sDate := DateFormat(stTime:= fbGetTime.dtDateAndTime);
//----------------------------------------------------------------------------------------------
// Delete
//----------------------------------------------------------------------------------------------
IF rtDelete.Q THEN
	FOR uiI := 1 TO cuiSize DO
		IF astErrorEvent[uiI].sErrorID = sErrorID THEN
			SysMemMove(pSrc := ADR(astErrorEvent[uiI+1]), pDest := ADR(astErrorEvent[uiI]), udiCount :=  SIZEOF(st_ErrorEvent) * (cuiSize-uiI));
			astErrorEvent[cuiSize].sErrorID		:= 'No error';
			EXIT;		
		END_IF
	END_FOR
END_IF

END_FUNCTION_BLOCK

// Programs/Tools/DateFormat
FUNCTION DateFormat : STRING
VAR_INPUT
	///Time input from ErrorFifo
	stTime: DATE_AND_TIME;
END_VAR
VAR
	///Date output in string
	sDate : STRING;
	sTemp : STRING;
	sDateTime: STRING := '';
END_VAR

//------------------------------------------------------------------------
// To show the date in the errortable in a usable format
//------------------------------------------------------------------------	

sDate := DT_TO_STRING(stTime);

//------------------------------------------------------------------------
// Cutting the days
//------------------------------------------------------------------------	

sTemp := sDate;
sDateTime := MID(STR:= sTemp, LEN:= 2, POS:= 12);
sDateTime := CONCAT(sDateTime, '/');
	
//------------------------------------------------------------------------
// Cutting the months
//------------------------------------------------------------------------		
sTemp := sDate;
sDateTime := CONCAT(sDateTime, MID(STR:= sTemp, LEN:= 2, POS:= 9));
sDateTime := CONCAT(sDateTime, '/');

//------------------------------------------------------------------------
// Cutting the years
//------------------------------------------------------------------------		

sTemp := sDate;
sDateTime := CONCAT(sDateTime, MID(STR:= sTemp, LEN:= 4, POS:= 4));
sDateTime := CONCAT(sDateTime, ' - ');	
	
//------------------------------------------------------------------------
// Cutting the hours and minutes and seconds
//------------------------------------------------------------------------	

sTemp := sDate;
sDateTime := CONCAT(sDateTime, RIGHT(STR:= sTemp, SIZE:= 8)	);

//------------------------------------------------------------------------		


	DateFormat := sDateTime;

END_FUNCTION

// Programs/Tools/MovCntr2B2M
FUNCTION_BLOCK MovCntr2B2M
VAR_INPUT
	/// Flag to Reset Error
	xQuit: BOOL;
	/// Enable error reset flag
	xQuitEN: BOOL;
	/// Enable error control
	xEnable: BOOL;
	/// Limit switch for movement 1 (M1 <--> B1) 
	xB1: BOOL;
	/// Limit switch for movement 2 (M2 <--> B2) 
	xB2: BOOL;
	/// Actor Signal for movement 1 (M1 <--> B1) 
	xM1: BOOL;
	/// Actor Signal for movement 1 (M2 <--> B2) 
	xM2: BOOL;
	/// Timeout-Time for movement 1	
	T1: TIME;
	/// Timeout-Time for movement 2
	T2: TIME;
END_VAR
VAR
	/// Timeout timer for movement 1
	TON1: TON;
	/// Timeout timer for movement 2
	TON2: TON;
	/// SR FlipFlop for Err1
	RS1: RS;
	/// SR FlipFlop for Err2
	RS2: RS;
END_VAR
VAR_OUTPUT
	/// Timeout movement 1
	xErr1: BOOL;
	/// Timeout movement 2 
	xErr2: BOOL;
END_VAR

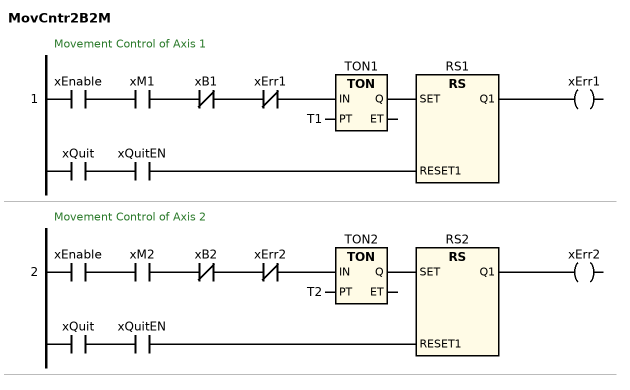
// NETWORK 1
// Movement Control of Axis 1
TON1(IN := xEnable AND xM1 AND NOT xB1 AND NOT xErr1, PT := T1); // TON
RS1(SET := TON1.Q, RESET1 := xQuit AND xQuitEN); // RS
xErr1 := RS1.Q1;

// NETWORK 2
// Movement Control of Axis 2
TON2(IN := xEnable AND xM2 AND NOT xB2 AND NOT xErr2, PT := T2); // TON
RS2(SET := TON2.Q, RESET1 := xQuit AND xQuitEN); // RS
xErr2 := RS2.Q1;

END_FUNCTION_BLOCK

// Programs/Visu/VisuProgramStp
PROGRAM  VisuProgramStp
VAR
	blBlink	: BLINK;
	t: TIME;
	uiNumOfApplications	: UINT:= 1;
	uiNumOfStoppers		: UINT:= 1;
	rtConvR				: R_TRIG;
	rtConvL				: R_TRIG;
	rtConvS				: R_TRIG;
	byActiveMainScreen	: BYTE;
	byActiveSubScreen	: BYTE;
	byScreenTitle		: BYTE;
	uiI					: UINT;
	astErrorEvents		: ARRAY [1..20] OF st_ErrorEvent;
	rtTime				: R_TRIG;
	fbGetTime: RTCLK.GetDateAndTime;
	sDate: STRING;
	dtTime	: DATE_AND_TIME;
	uiCarrierInitNum: UINT;
	xCarrierInit: BOOL;
	tonDefErr: TON;
	tonMesErr: TON;
	tonSapErr: TON;
	
	stRfidCdpx	: dc_ecp.st_CPF_RfidData;
	astAppControlONo: UDINT;
END_VAR

byActiveMainScreen	:= BOOL_TO_BYTE(fromCDPX.stCdpxButtonState.xHome)*0 + BOOL_TO_BYTE(fromCDPX.stCdpxButtonState.xSetupMode)*1 + BOOL_TO_BYTE(fromCDPX.stCdpxButtonState.xParameter)*2 + BOOL_TO_BYTE(fromCDPX.stCdpxButtonState.xSystem)*3;
byActiveSubScreen	:= BOOL_TO_BYTE(fromCDPX.stCdpxButtonState.xOperationMode)*0 + BOOL_TO_BYTE(fromCDPX.stCdpxButtonState.xApp_1)*0 +  BOOL_TO_BYTE(fromCDPX.stCdpxButtonState.xApp)*0 + BOOL_TO_BYTE(fromCDPX.stCdpxButtonState.xSystem)*0 + BOOL_TO_BYTE(fromCDPX.stCdpxButtonState.xOverview)*1 + BOOL_TO_BYTE(fromCDPX.stCdpxButtonState.xApp_2)*1 +  BOOL_TO_BYTE(fromCDPX.stCdpxButtonState.xTrans_1)*1 + BOOL_TO_BYTE(fromCDPX.stCdpxButtonState.xUser)*2 + BOOL_TO_BYTE(fromCDPX.stCdpxButtonState.xBelt)*2 +  BOOL_TO_BYTE(fromCDPX.stCdpxButtonState.xTrans_2)*2 + BOOL_TO_BYTE(fromCDPX.stCdpxButtonState.xStp_1)*3+ BOOL_TO_BYTE(fromCDPX.stCdpxButtonState.xStp_2)*4;
byScreenTitle 		:= byActiveMainScreen* 10 + byActiveSubScreen  ;

dtTime := fbGetTime.dtDateAndTime;
rtTime(CLK:= fbGetTime.xDone);
IF rtTime.Q THEN
sDate := DateFormat(stTime:= dtTime);
END_IF
fbGetTime( xExecute:= NOT fbGetTime.xDone);
fbGetTime( xExecute:= fbGetTime.xDone);

//////////////////////////////////
//			from CDPX			//
//////////////////////////////////

IF xFirstCycle THEN
	fromCDPX.astTransitionTable_1:= astTransitionTableStopper1 ;
	fromCDPX.uiMode := 1;
ELSE	
	astTransitionTableStopper1 :=fromCDPX.astTransitionTable_1;
	Visu.byMode 			:= UINT_TO_BYTE(fromCDPX.uiMode);
END_IF

// DABO /////////////////////////////////////////////////////////////////////////
IF uiCarrierInitNum <> stpStopper1.stAppSettings.uiCarrierInitNum THEN
	uiCarrierInitNum := stpStopper1.stAppSettings.uiCarrierInitNum;
ELSIF uiCarrierInitNum <> fromCDPX.astAppSetting[0].uiCarrierInitNum THEN
	uiCarrierInitNum := fromCDPX.astAppSetting[0].uiCarrierInitNum;
END_IF

fromCDPX.astAppSetting[0].uiCarrierInitNum := uiCarrierInitNum;
SysMemCpy(pDest:= ADR(stpStopper1.stAppSettings.uiCarrierInitNum), pSrc:= ADR(uiCarrierInitNum), udiCount:= SIZEOF(uiCarrierInitNum));

IF xCarrierInit <> stpStopper1.stAppSettings.xCarrierInit THEN
	xCarrierInit := stpStopper1.stAppSettings.xCarrierInit;
ELSIF xCarrierInit <> fromCDPX.astAppSetting[0].xCarrierInit THEN
	xCarrierInit := fromCDPX.astAppSetting[0].xCarrierInit;
END_IF

fromCDPX.astAppSetting[0].xCarrierInit := xCarrierInit;
SysMemCpy(pDest:= ADR(stpStopper1.stAppSettings.xCarrierInit), pSrc:= ADR(xCarrierInit), udiCount:= SIZEOF(xCarrierInit));

SysMemCpy(pDest:= ADR(stpStopper1.stAppSettings.xActive), pSrc:= ADR(fromCDPX.astAppSetting[0].xActive), udiCount:= SIZEOF(fromCDPX.astAppSetting[0].xActive));
SysMemCpy(pDest:= ADR(stpStopper1.stAppSettings.xStopBelt), pSrc:= ADR(fromCDPX.astAppSetting[0].xStopBelt), udiCount:= SIZEOF(fromCDPX.astAppSetting[0].xStopBelt));

//////////////////////////////////////////////////////////////////////////////////
// conveyor handling
rtConvL(CLK:= fromCDPX.astConveyorButtonState[0].xConvLeft);
rtConvR(CLK:= fromCDPX.astConveyorButtonState[0].xConvRight);
rtConvS(CLK:= fromCDPX.astConveyorButtonState[0].xConvSlow);
IF rtConvL.Q THEN
	IF  stpStopper1.convConveyor.xLeft THEN
		stpStopper1.convConveyor.Stop();
	ELSE
		stpStopper1.convConveyor.RunToLeft(stpStopper1.convConveyor.xSlow);
	END_IF
END_IF
IF rtConvR.Q THEN
	IF  stpStopper1.convConveyor.xRight THEN
		stpStopper1.convConveyor.Stop();
	ELSE
		stpStopper1.convConveyor.RunToRight(stpStopper1.convConveyor.xSlow);
	END_IF
END_IF
IF rtConvS.Q THEN
	IF  stpStopper1.convConveyor.xSlow THEN
		stpStopper1.convConveyor.SpeedUp();
	ELSE
		stpStopper1.convConveyor.SlowDown();
	END_IF
END_IF

// Operation mode buttons
fromCDPX.stHome_OperationMode_Reset.xActive := xReset OR (xResetEn AND blBlink.OUT);
fromCDPX.stHome_OperationMode_Reset.xDisabled := NOT xResetEn;

fromCDPX.stHome_OperationMode_Automatic.xActive := xAuto OR (xAutoEn AND blBlink.OUT);
fromCDPX.stHome_OperationMode_Automatic.xDisabled := NOT xAutoEn AND NOT xAuto;

fromCDPX.stHome_OperationMode_Setup.xActive := xManual;
fromCDPX.stHome_OperationMode_Setup.xDisabled := NOT xManualEn AND NOT xManual;

fromCDPX.stHome_OperationMode_CycleEnd.xActive := xCycleEnd AND blBlink.OUT;
fromCDPX.stHome_OperationMode_CycleEnd.xDisabled := NOT xCycleEndEn AND NOT xCycleEnd;

stWinCC.xAuto 		:= fromCDPX.stHome_OperationMode_Automatic.xPressed;
stWinCC.xReset 		:= fromCDPX.stHome_OperationMode_Reset.xPressed;
stWinCC.xManual 	:= fromCDPX.stHome_OperationMode_Setup.xPressed;
stWinCC.xCycleEnd 	:= fromCDPX.stHome_OperationMode_CycleEnd.xPressed;
stWinCC.xQuit		:= fromCDPX.stCdpxButtonState.xClearError;

// Setup RFID buttons
fromCDPX.stSetupMode_Stopper1_Init.xActive R= stpStopper1.stpStopper.dtmRfid.xReady;
fromCDPX.stSetupMode_Stopper1_Init.xActive S= fromCDPX.stSetupMode_Stopper1_Init.xPressed;
fromCDPX.stSetupMode_Stopper1_Init.xDisabled :=  xManual;
IF fromCDPX.astStopperButton[0].xInit THEN
	stpStopper1.stpStopper.Connect(usiCanChannel := stpStopper1.usiCanChannel, usiCanNetworkId := stpStopper1.usiCanNetworkId, usiCanNodeId := stpStopper1.usiCanNodeId);
END_IF


fromCDPX.stSetupMode_Stopper1_Read.xActive R= stpStopper1.stpStopper.dtmRfid.xReady;
fromCDPX.stSetupMode_Stopper1_Read.xActive S= fromCDPX.stSetupMode_Stopper1_Read.xPressed;
fromCDPX.stSetupMode_Stopper1_Read.xDisabled := xManual;
IF fromCDPX.astStopperButton[0].xRead THEN
	stpStopper1.stpStopper.ReadRfid(pstRfidData := ADR(stRfidCdpx));
	toCDPX.astRfidData[0].uiCarrierID				:=	stRfidCdpx.uiCarrierID					 ;
	toCDPX.astRfidData[0].uiCode					:=	stRfidCdpx.uiCode						 	;
	toCDPX.astRfidData[0].uiParameter1				:=	stRfidCdpx.uiParameter1					 ;
	toCDPX.astRfidData[0].uiParameter2				:=	stRfidCdpx.uiParameter2					 ;
	toCDPX.astRfidData[0].uiParameter3				:=	stRfidCdpx.uiParameter3					 ;
	toCDPX.astRfidData[0].uiParameter4				:=	stRfidCdpx.uiParameter4					 ;
	toCDPX.astRfidData[0].stMesData.udiONo			:=	stRfidCdpx.stMesData.udiONo				 ;
	toCDPX.astRfidData[0].stMesData.udiPNo			:=	stRfidCdpx.stMesData.udiPNo				 ;
	toCDPX.astRfidData[0].stMesData.uiOpNo			:=	stRfidCdpx.stMesData.uiOpNo				 ;
	toCDPX.astRfidData[0].stMesData.uiOPos			:=	stRfidCdpx.stMesData.uiOPos				 ;
	toCDPX.astRfidData[0].stMesData.uiResourceId	:=	stRfidCdpx.stMesData.uiResourceId		 	;
	toCDPX.astRfidData[0].stSapData.sItem	 		:=	stRfidCdpx.stSapData.sItem	 			 ;
	toCDPX.astRfidData[0].stSapData.sItemRev		:=	stRfidCdpx.stSapData.sItemRev			 	;
	toCDPX.astRfidData[0].stSapData.sSfc			:=	stRfidCdpx.stSapData.sSfc				 	;
	toCDPX.astRfidData[0].stSapData.udiOp			:=	stRfidCdpx.stSapData.udiOp				 ;
	toCDPX.astRfidData[0].stSapData.udiSfc			:=	stRfidCdpx.stSapData.udiSfc				 ;
END_IF                                                	


fromCDPX.stSetupMode_Stopper1_Write.xActive R= stpStopper1.stpStopper.dtmRfid.xReady;
fromCDPX.stSetupMode_Stopper1_Write.xActive S= fromCDPX.stSetupMode_Stopper1_Write.xPressed;
fromCDPX.stSetupMode_Stopper1_Write.xDisabled := xManual;
IF fromCDPX.astStopperButton[0].xWrite THEN
	stRfidCdpx.uiCarrierID					:= toCDPX.astRfidData[0].uiCarrierID				;
	stRfidCdpx.uiCode						:= toCDPX.astRfidData[0].uiCode					;
	stRfidCdpx.uiParameter1					:= toCDPX.astRfidData[0].uiParameter1				;
	stRfidCdpx.uiParameter2					:= toCDPX.astRfidData[0].uiParameter2				;
	stRfidCdpx.uiParameter3					:= toCDPX.astRfidData[0].uiParameter3				;
	stRfidCdpx.uiParameter4					:= toCDPX.astRfidData[0].uiParameter4				;
	stRfidCdpx.stMesData.udiONo				:= toCDPX.astRfidData[0].stMesData.udiONo			;
	stRfidCdpx.stMesData.udiPNo				:= toCDPX.astRfidData[0].stMesData.udiPNo			;
	stRfidCdpx.stMesData.uiOpNo				:= toCDPX.astRfidData[0].stMesData.uiOpNo			;
	stRfidCdpx.stMesData.uiOPos				:= toCDPX.astRfidData[0].stMesData.uiOPos			;
	stRfidCdpx.stMesData.uiResourceId		:= toCDPX.astRfidData[0].stMesData.uiResourceId	;
	stRfidCdpx.stSapData.sItem	 			:= toCDPX.astRfidData[0].stSapData.sItem	 		;
	stRfidCdpx.stSapData.sItemRev			:= toCDPX.astRfidData[0].stSapData.sItemRev		;
	stRfidCdpx.stSapData.sSfc				:= toCDPX.astRfidData[0].stSapData.sSfc			;
	stRfidCdpx.stSapData.udiOp				:= toCDPX.astRfidData[0].stSapData.udiOp			;
	stRfidCdpx.stSapData.udiSfc				:= toCDPX.astRfidData[0].stSapData.udiSfc			;
	stpStopper1.stpStopper.WriteRfid(stRfidData:= stRfidCdpx);
END_IF


fromCDPX.stSetupMode_Stopper1_DeleteData.xActive := fromCDPX.stSetupMode_Stopper1_DeleteData.xPressed;
fromCDPX.stSetupMode_Stopper1_DeleteData.xDisabled := xManual;                                            
IF fromCDPX.astStopperButton[0].xDeleteData	THEN
	SysMemSet(pDest:= ADR(stpStopper1.stpStopper.stRfidVisu), udiValue:= 0, udiCount:= SIZEOF(stpStopper1.stpStopper.stRfidVisu));
	SysMemCpy(pDest:= ADR(toCDPX.astRfidData[0]), pSrc:= ADR(stpStopper1.stpStopper.stRfidVisu), udiCount:= SIZEOF(stpStopper1.stpStopper.stRfidData));	
END_IF

IF NOt xManual  THEN
	SysMemCpy(pDest:= ADR(toCDPX.astRfidData[0]), pSrc:= ADR(stpStopper1.stpStopper.stRfidVisu), udiCount:= SIZEOF(stpStopper1.stpStopper.stRfidData));	
END_IF


IF fromCDPX.astStopperButton[0].xStpMveDown	THEN
	stpStopper1.stpStopper.cpfssStopper.StayDown();
END_IF
IF fromCDPX.astStopperButton[0].xStpMveUp	THEN
	stpStopper1.stpStopper.cpfssStopper.MoveUp();
END_IF

Visu.stInteractiveError.xBtnAbort 		:= fromCDPX.stInteractiveMessage_Abort.xPressed;
Visu.stInteractiveError.xBtnIgnore 		:= fromCDPX.stInteractiveMessage_Ignore.xPressed;
Visu.stInteractiveError.xBtnRejectOrder := fromCDPX.stInteractiveMessage_RejectOrder.xPressed;
Visu.stInteractiveError.xBtnRepeat		:= fromCDPX.stInteractiveMessage_Repeat.xPressed;

blBlink(ENABLE := TRUE, TIMEHIGH := T#1S, TIMELOW := T#1S); 
	

IF Visu.byMode = 1 THEN
	xMES := TRUE;
	xSAP := FALSE;
ELSIF Visu.byMode = 2 THEN
	xMES := FALSE;
	xSAP := TRUE;
ELSE
	xMES := FALSE;
	xSAP := FALSE;
END_IF

IF NOT xAuto AND NOT xManual AND NOT xReset THEN
	Visu.byOpMode := 0;
ELSIF xReset THEN
	Visu.byOpMode := 1;
ELSIF xAuto THEN
	Visu.byOpMode := 2;
ELSIF xManual THEN
	Visu.byOpMode := 3;
END_IF


//////////////////////////////////
//			to CDPX				//
//////////////////////////////////


toCDPX.byOpMode									:= Visu.byOpMode;
toCDPX.byScreenTitle							:= byScreenTitle;
toCDPX.xManual									:= xManual;	
toCDPX.xAuto									:= xAuto;			
toCDPX.xSAP										:= xSAP;				
toCDPX.xMES										:= xMES;				
toCDPX.xDefault									:= NOT xSAP AND NOT xMES;		
toCDPX.uiNumOfApplications						:= uiNumOfApplications;				
toCDPX.uiNumOfStoppers							:= uiNumOfStoppers;						
toCDPX.sDate									:= LEFT(sDate,10);
toCDPX.sTime									:= RIGHT(sDate,8);
toCDPX.auiCondIn[0]								:= stpStopper1.uiCondIn;
toCDPX.auiCondOut[0]							:= stpStopper1.uiCondOut;


toCDPX.astSensorSignals[0].sInductive_1			:= 'xBG21';
toCDPX.astSensorSignals[0].sInductive_2			:= 'xBG22';
toCDPX.astSensorSignals[0].sInductive_3			:= 'xBG23';
toCDPX.astSensorSignals[0].sInductive_4			:= 'xBG24';
toCDPX.astSensorSignals[0].sRfid				:= 'TF80';
toCDPX.astSensorSignals[0].sStpDownOutpu		:= 'xMB20';
toCDPX.astSensorSignals[0].sStpDownSensor		:= 'xBG20';
toCDPX.astSensorSignals[0].xInductive_1			:= xBG21; 
toCDPX.astSensorSignals[0].xInductive_2			:= xBG22; 
toCDPX.astSensorSignals[0].xInductive_3			:= xBG23; 
toCDPX.astSensorSignals[0].xInductive_4			:= xBG24; 
toCDPX.astSensorSignals[0].xStpDownOutpu		:= xMB20; 
toCDPX.astSensorSignals[0].xStpDownSensor		:= xBG20;
toCDPX.astSensorSignals[0].xTagPresent			:= stpStopper1.stpStopper.dtmRfid.stState.xTagPresent;
toCDPX.astSensorSignals[0].xReady				:= stpStopper1.stpStopper.dtmRfid.xReady;
toCDPX.astSensorSignals[0].xBusy				:= NOT stpStopper1.stpStopper.dtmRfid.xReady;
toCDPX.astSensorSignals[0].xError				:= stpStopper1.stpStopper.dtmRfid.xError;
toCDPX.astSensorSignals[0].xTimeOut				:= stpStopper1.stpStopper.dtmRfid.xTimeout;
                                               
toCDPX.astConveyorSignals[0].sConvLeft			:= 'QA1_R';
toCDPX.astConveyorSignals[0].sConvRight			:= 'QA1_L';
toCDPX.astConveyorSignals[0].sConvSlow			:= 'QA1_S';
toCDPX.astConveyorSignals[0].xConvMovingLeft	:= stpStopper1.convConveyor.xLeft;
toCDPX.astConveyorSignals[0].xConvMovingRight	:= stpStopper1.convConveyor.xRight;
toCDPX.astConveyorSignals[0].xConvMovingSlow	:= stpStopper1.convConveyor.xSlow;

toCDPX.astAppState[0] 		:= stpStopper1.stAppState;
toCDPX.astAppControl[0]		:= AppModul.stAppControl;
astErrorEvents				:= Visu.fbErrorFifo.astErrorEvent;

tonDefErr(IN := Visu.stInteractiveError.xError AND NOT xMES AND NOT xSAP, PT := T#0.5S);
tonMesErr(IN := Visu.stInteractiveError.xError AND (xMES OR (xSAP AND stpStopper1.uiState <> 999)), PT := T#0.5S);
tonSapErr(IN := Visu.stInteractiveError.xError AND NOT xMES AND xSAP AND stpStopper1.uiState = 999, PT := T#0.5S);


toCDPX.stInteractiveErrors.uiIntMsgID	:= STRING_TO_UINT(Visu.stInteractiveError.sMessageID);
toCDPX.stInteractiveErrors.xIntDefault	:= tonDefErr.Q;
toCDPX.stInteractiveErrors.xIntMES		:= tonMesErr.Q;
toCDPX.stInteractiveErrors.xIntSAP		:= tonSapErr.Q;
toCDPX.stInteractiveErrors.uiIntAbort	:= Visu.stInteractiveError.uiAbortState;
toCDPX.stInteractiveErrors.uiIntIgnore	:= Visu.stInteractiveError.uiIgnoreState;
toCDPX.stInteractiveErrors.uiIntState	:= Visu.stInteractiveError.uiState;
toCDPX.stInteractiveErrors.sSapError	:= SAPHMI.sError;
toCDPX.stInteractiveErrors.udiSapSfc	:= SAPHMI.udiSfc;
toCDPX.stInteractiveErrors.uiSapOp		:= SAPHMI.uiOp;
toCDPX.stInteractiveErrors.uiSapPos		:= SAPHMI.uiPos;

FOR uiI := 1 TO 20 DO
	IF astErrorEvents[uiI].sErrorID <> 'No error' THEN
		toCDPX.astErrors[uiI].xError := TRUE;
		toCDPX.astErrors[uiI].uiLevel			:= STRING_TO_UINT(RIGHT(LEFT(astErrorEvents[uiI].sErrorID,2),1))+1;
		toCDPX.astErrors[uiI].uiMsgNum			:= toCDPX.astErrors[uiI].uiLevel*10 + STRING_TO_UINT(RIGHT(astErrorEvents[uiI].sErrorID,1));
 		toCDPX.astErrors[uiI].sErrorID			:= astErrorEvents[uiI].sErrorID;
		toCDPX.astErrors[uiI].sDateTime			:= astErrorEvents[uiI].sDateTime;
	ELSE                                		
		toCDPX.astErrors[uiI].xError 			:= FALSE;
		toCDPX.astErrors[uiI].uiLevel			:= 0;
		toCDPX.astErrors[uiI].uiMsgNum			:= 0;
		toCDPX.astErrors[uiI].sErrorID			:= '';
		toCDPX.astErrors[uiI].sDateTime			:= '';
	END_IF	
END_FOR

toCDPX.auiCarrierInitNum[0]	:= stpStopper1.uiCarrierInitNum;

//SysMemCpy(pDest:= ADR(), pSrc:= ADR(), udiCount:= SIZEOF());

END_PROGRAM

// Programs/TrafficStopper
FUNCTION_BLOCK TrafficStopper
VAR_INPUT
	xCarrierAvSensor: BOOL;
	xStopperReleased: BOOL;
	xSemaIn			: BOOL;
END_VAR
VAR_OUTPUT
	xInitPos			: BOOL;
	xLeft				: BOOL;
	xRight				: BOOL;
	xSlow				: BOOL;
	xStop				: BOOL;
	xReleaseStopper		: BOOL;
	xSemaOut			: BOOL;
END_VAR
VAR
	uiState				: UINT := 0;
	convConveyor		: dc_ecp.Conveyor2Dir;
	stpStopper			: dc_ecp.CPF_StopperSimple;
	ftAuto				: F_TRIG;
	ftManual			: F_TRIG;
	uiNextState: UINT;
	uiI: UINT;
	uiCondIn		: UINT;
	uiCondOut		: UINT;

END_VAR

xSemaOut := xSemaIn;

////////////////////////////////////////////
// Execute moduls
////////////////////////////////////////////

_ModuleCalls();

////////////////////////////////////////////
// Exit from auto or manual mode
////////////////////////////////////////////

ftAuto(CLK := xAuto);
ftManual(CLK := xManual);

IF ftAuto.Q OR ftManual.Q THEN
	convConveyor.Stop();
	stpStopper.MoveUp();
	uiState := 0;
END_IF

xInitPos := (uiState <= 10);


////////////////////////////////////////////
// Default Mode
////////////////////////////////////////////

// Execute Default Mode
IF xAuto THEN
	_DefaultMode();
END_IF

METHOD PRIVATE _DefaultMode : BOOL
VAR_INPUT
END_VAR
CASE uiState OF
	0:	// Idle
		convConveyor.Stop();
		IF xAuto THEN
			uiState := 1;
		END_IF
		
	1:	// Init
		convConveyor.RunToRight(FALSE);
		uiState := 2;
		
	
	2:	// Wait for RFID
		IF stpStopper.xReady  THEN
			uiState := 10;
		END_IF
		
	10:	// Wait until carrier at stopper
		IF stpStopper.xCarrierAvailable AND NOT xCycleEnd THEN
			uiState := 500;
		END_IF
		
	500:// Pass carrier
		IF NOT xSemaIn THEN
			xSemaOut := TRUE;
			stpStopper.Release();
			uiState := 505;
		END_IF
		
	505:// Wait for release
		IF stpStopper.xReady THEN
			uiState := 10;
		END_IF
	
END_CASE
END_METHOD

METHOD PRIVATE _ModuleCalls : BOOL
VAR_INPUT
END_VAR
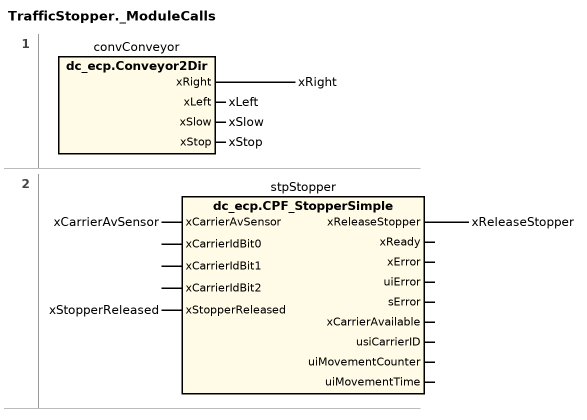
// NETWORK 1
convConveyor(xLeft => xLeft, xSlow => xSlow, xStop => xStop); // dc_ecp.Conveyor2Dir
xRight := convConveyor.xRight;

// NETWORK 2
stpStopper(xCarrierAvSensor := xCarrierAvSensor, xStopperReleased := xStopperReleased); // dc_ecp.CPF_StopperSimple
xReleaseStopper := stpStopper.xReleaseStopper;
END_METHOD

END_FUNCTION_BLOCK

// Programs/Tools/MovCntr3B3M
FUNCTION_BLOCK MovCntr3B3M
VAR_INPUT
	/// Flag to Reset Error
	xQuit: BOOL;
	/// Enable error reset flag
	xQuitEN: BOOL;
	/// Enable error control
	xEnable: BOOL;
	/// Limit switch for movement 1 (M1 <--> B1) 
	xB1: BOOL;
	/// Limit switch for movement 2 (M2 <--> B2) 
	xB2: BOOL;
	/// Limit switch for movement 2 (M3 <--> B3) 
	xB3: BOOL;
	/// Actor Signal for movement 1 (M1 <--> B1)
	xM1: BOOL;
	/// Actor Signal for movement 1 (M2 <--> B2)
	xM2: BOOL;
	/// Actor Signal for movement 1 (M3 <--> B3) 
	xM3: BOOL;
	/// Timeout-Time for movement 1	
	T1: TIME;
	/// Timeout-Time for movement 2
	T2: TIME;
	/// Timeout-Time for movement 3	
	T3: TIME;
END_VAR
VAR
	/// Timeout timer for movement 1
	TON1: TON;
	/// Timeout timer for movement 2
	TON2: TON;
	/// Timeout timer for movement 3
	TON3: TON;
	/// SR FlipFlop for Err1
	SR1: SR;
	/// SR FlipFlop for Err2
	SR2: SR;
	/// SR FlipFlop for Err3
	SR3: SR;
END_VAR
VAR_OUTPUT
	/// Timeout movement 1 
	xErr1: BOOL;
	/// Timeout movement 2 
	xErr2: BOOL;
	/// Timeout movement 3 
	xErr3: BOOL;
END_VAR

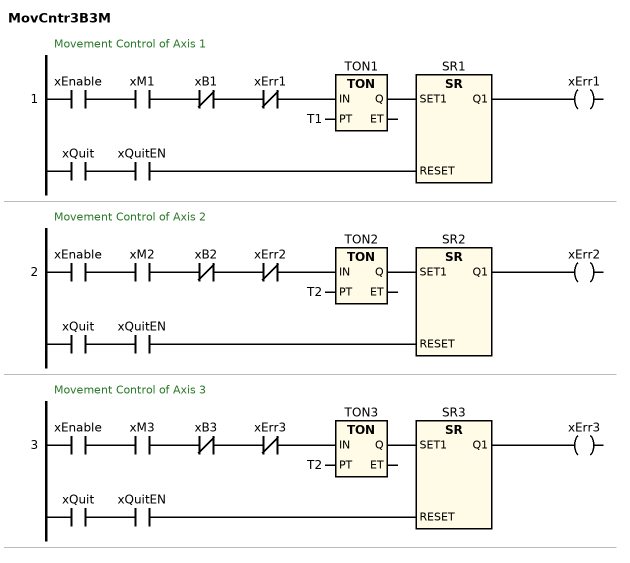
// NETWORK 1
// Movement Control of Axis 1
TON1(IN := xEnable AND xM1 AND NOT xB1 AND NOT xErr1, PT := T1); // TON
SR1(SET1 := TON1.Q, RESET := xQuit AND xQuitEN); // SR
xErr1 := SR1.Q1;

// NETWORK 2
// Movement Control of Axis 2
TON2(IN := xEnable AND xM2 AND NOT xB2 AND NOT xErr2, PT := T2); // TON
SR2(SET1 := TON2.Q, RESET := xQuit AND xQuitEN); // SR
xErr2 := SR2.Q1;

// NETWORK 3
// Movement Control of Axis 3
TON3(IN := xEnable AND xM3 AND NOT xB3 AND NOT xErr3, PT := T2); // TON
SR3(SET1 := TON3.Q, RESET := xQuit AND xQuitEN); // SR
xErr3 := SR3.Q1;

END_FUNCTION_BLOCK

// Programs/StopperWithMes
FUNCTION_BLOCK StopperWithMes
VAR_INPUT
	byMode				: BYTE;
	usiCanNodeId		: USINT := 32;
	usiCanNetworkId		: USINT := 0;
	usiCanChannel		: USINT := 1;
	sMesIp				: STRING := '172.20.0.90';
	uiMesQueryPort		: UINT := 2000;
	uiMesStatePort		: UINT := 2001;
	uiResourceId		: UINT := 0;
	stAppState			: st_AppState;
	stAppInfo			: st_AppInfo;
	xFirstSapModule		: BOOL	:= FALSE;
	udiMyOp				: UDINT;

	xRfid_SiemensByteOrder: BOOL;
	xCarrierAvSensor: BOOL;
	xCarrierIdBit0: BOOL;
	xCarrierIdBit1: BOOL;
	xCarrierIdBit2: BOOL;
	xStopperReleased: BOOL;
	xSemaIn			: BOOL;
	xParametricData	:BOOL;
	
	
END_VAR
VAR_OUTPUT
	xInitPos			: BOOL;
	xLeft				: BOOL;
	xRight				: BOOL;
	xSlow				: BOOL;
	xStop				: BOOL;
	stAppControl		: st_AppControl;
	stAppSettings		: st_AppSettings;

	xReleaseStopper		: BOOL;
	xSemaOut			: BOOL;
END_VAR
VAR_IN_OUT
	astTransitionTable	: ARRAY [0..10] OF st_TransitionData;
END_VAR
VAR
	uiState				: UINT := 0;
	convConveyor		: dc_ecp.Conveyor2Dir;
	stpStopper			: dc_ecp.CPF_StopperDtm425;
	mesMES				: dc_ecp.MES4;
	stRfidData			: dc_ecp.st_CPF_RfidData;
	stRcvHeader			: dc_ecp.st_MES4_QueryHeader;
	auiRcvPar			: ARRAY [0..3] OF UINT;
	auiSndPar			: ARRAY [0..3] OF UINT;
	xFirstWorkOrder		: BOOL := FALSE;
	udiONo				: UDINT;
	uiOPos				: UINT;
	uiOpNo				: UINT;
	uiCarrierId			: UINT;
	ftAuto				: F_TRIG;
	ftManual			: F_TRIG;
	uiActualTransitionRow: UINT;
	uiNextState: UINT;
	uiI: UINT;
	xValidOperation: BOOL;
	uiCarrierInitNum	: UINT;
	uiCondIn		: UINT;
	uiCondOut		: UINT;

	// SAP //
	uiErrNo: UINT;
	udiSfc           : UDINT;
    udiOp            : UDINT;	
	tonHs: TON;
	tonOpc: TON;	
	abySapParameter : ARRAY [0..3] OF INT;
	tTimeOutHs		: TIME := T#5S;
	uiRetryState	: UINT;	
		
	tonMES: TON;
END_VAR

xSemaOut := xSemaIn;

////////////////////////////////////////////
// Execute moduls
////////////////////////////////////////////

_ModuleCalls();

		
////////////////////////////////////////////
// Init RFID
////////////////////////////////////////////
IF NOT stpStopper.xConnected AND stpStopper.xReady THEN	
	stpStopper.Connect(usiCanNodeId:= usiCanNodeId, usiCanNetworkId:= usiCanNetworkId, usiCanChannel:= usiCanChannel);
END_IF

////////////////////////////////////////////
// MES Mode
////////////////////////////////////////////

// Execute MES mode
IF xAuto AND byMode = 1 THEN
	_MesMode();
END_IF

// Connect to MES
IF NOT mesMES.xConnected AND mesMES.xReady OR mesMES.xError THEN
	mesMES.Connect(sIP := sMesIp, uiQueryPort := uiMesQueryPort, uiStatePort := uiMesStatePort, uiResourceId := uiResourceId);
END_IF


////////////////////////////////////////////
// Exit from auto or manual mode
////////////////////////////////////////////

ftAuto(CLK := xAuto);
ftManual(CLK := xManual);

IF ftAuto.Q OR ftManual.Q THEN
	convConveyor.Stop();
	stpStopper.cpfssStopper.MoveUp();
	uiState := 0;
END_IF

stAppControl.xReset := xReset;

mesMES.stResourceState.xAuto := xAuto;
mesMES.stResourceState.xManual := xManual;
mesMES.stResourceState.xReset := xReset;
mesMES.stResourceState.xMES := xMES;
mesMES.stResourceState.xErrL0 := stError.xSF0;
mesMES.stResourceState.xErrL1 := stError.xSF1;
mesMES.stResourceState.xErrL2 := stError.xSF2;
mesMES.stResourceState.xBusy := NOT stAppState.xReady;

xInitPos := (uiState <= 10) AND (stAppState.xInitPos OR NOT stAppSettings.xActive);


////////////////////////////////////////////
// Default Mode
////////////////////////////////////////////

// Execute Default Mode
IF xAuto AND byMode = 0 THEN
	_DefaultMode();
END_IF

////////////////////////////////////////////
// SAP Mode
////////////////////////////////////////////

// Execute SAP Mode
IF xAuto AND byMode = 2 THEN
	_SapMode(xFirstSapModule := xFirstSapModule, udiMyOp := udiMyOp);
END_IF

METHOD PRIVATE _MesMode : BOOL
VAR_INPUT
END_VAR

VAR
	uiErrNo: UINT;
END_VAR
CASE uiState OF
	0:	// Idle
		convConveyor.Stop();
		IF xAuto THEN
			uiState := 1;
		END_IF		
	
	1: // Init
		IF mesMES.xConnected THEN
			convConveyor.RunToRight(FALSE);
			uiState := 2;
		END_IF	
		
		
	2:	// Wait for RFID
		IF stpStopper.xReady AND stpStopper.xConnected THEN
			uiState := 10;
		END_IF
	
		
	10:	// Wait until carrier at stopper
		IF stpStopper.xCarrierAvailable AND NOT xCycleEnd  THEN
			uiState := 15;
		END_IF
		
	15:	// Check if RFID tag recognized
		IF stpStopper.dtmRfid.stState.xTagPresent THEN
			uiState := 20;
		ELSE
			uiState := 500;
		END_IF
		
	20:	// Read RFID
		stpStopper.ReadRfid(ADR(stRfidData));
		uiState := 25;
		
	25:	// Wait until read finished
		IF stpStopper.xReady THEN
			uiCarrierId := stRfidData.uiCarrierID;
			uiState := 100;
		END_IF
		
	100:// App. ready and active?
		IF stAppState.xReady AND stAppSettings.xActive THEN
			uiState := 105;
		ELSE
			uiState := 500;
		END_IF
		
	105:// Carrier already asigned?
		IF stRfidData.stMesData.udiONo <> 0 AND stRfidData.stMesData.uiOPos <> 0 THEN
			uiState := 110;
		ELSE
			uiState := 115;
		END_IF
		
	110:// Get this order
		xFirstWorkOrder := FALSE;
		mesMES.GetOpForONoOPos(udiONo := stRfidData.stMesData.udiONo, uiOPos := stRfidData.stMesData.uiOPos, pRcvHeader := ADR(stRcvHeader), pRcvPar := ADR(auiRcvPar), szRcvPar := SIZEOF(auiRcvPar));
		uiState := 120;
		
	115:// Get order for resource
		xFirstWorkOrder := TRUE;
		mesMES.GetFirstOpForRsc(uiResourceId := uiResourceId, pRcvHeader := ADR(stRcvHeader), pRcvPar := ADR(auiRcvPar), szRcvPar := SIZEOF(auiRcvPar));
		uiState := 120;

	120:// Wait for MES request
		IF stRcvHeader.xDone THEN
			udiONo := strcvHeader.udiONo;
		    uiOPos := strcvHeader.uiOPos;
		    uiOpNo := strcvHeader.uiOpNo;
			uiState := 125;
		ELSIF xCycleEnd THEN
			uiState := 500;	
		END_IF

	125:// Order Available?
		IF udiONo <> 0 AND uiOPos <> 0 AND strcvHeader.uiResourceId = uiResourceId THEN
			uiState := 130;
		ELSE
			uiState := 135;
		END_IF	

	130:// Operation number is good?
		xValidOperation := FALSE;
		IF stAppInfo.byNumberOfOperations > 0 THEN
			FOR uiI := 0 TO stAppInfo.byNumberOfOperations - 1 DO
				IF stAppInfo.auiOperations[uiI] = uiOpNo THEN
					xValidOperation := TRUE;
					EXIT;
				END_IF
			END_FOR
		END_IF
	
		IF xValidOperation THEN
			uiState := 300;
		ELSE
			uiState := 500;
		END_IF
		
	135:// First Work Order?
		IF xFirstWorkOrder THEN
			uiState := 500;
		ELSE
			uiState := 400;
		END_IF
		
	300:// Wait app. free
		IF stAppSettings.xActive AND stAppState.xReady THEN
			uiState := 305;
		END_IF
		
	305:// Send parameters to app
		stAppControl.udiONo := udiONo;
		stAppControl.uiOPos := uiOPos;
		stAppControl.uiOpNo := uiOpNo;
		stAppControl.auiPar := auiRcvPar;
		toCDPX.astAppControlONo	:= udiONo;
		uiState := 310;
		
	310:// Send Start (OPStart)
		mesMES.OpStart(udiONo := udiONo, uiOPos := uiOPos, pRcvHeader := ADR(stRcvHeader));
		uiState := 320;
		
	320:// Wait for MES request
		IF stRcvHeader.xDone THEN
			uiState := 325;
		END_IF
		
	325:// Trigger App. start
		IF stAppSettings.xStopBelt THEN
			convConveyor.Stop();
		END_IF
		stAppControl.xStart := TRUE;
		uiState := 328;
		
	328:// Wait for App. started	
		IF NOT stAppState.xReady THEN
			stAppControl.xStart := FALSE;
			uiState := 330;
		END_IF
		
	330:// Wait for App. finished
		IF stAppState.xReady THEN
			convConveyor.RunToRight(FALSE);
			toCDPX.astAppControlONo	:= 0;
			uiState := 335;
		END_IF
		
	335:// App. fininshed without error?
		IF stAppState.uiReturnCode = 0 THEN
			uiState := 340;
		ELSE
			uiState := 336;
		END_IF
		
	336:// Interactive message
		Visu.stInteractiveError.xError := TRUE;
		Visu.stInteractiveError.sMessageID := UINT_TO_STRING(stAppState.uiReturnCode);
		visu.stInteractiveError.uiAbortState := 340;
		visu.stInteractiveError.uiIgnoreState := 340;
		
		// Retry
		IF visu.stInteractiveError.xBtnRepeat THEN
			visu.stInteractiveError.xBtnRepeat := FALSE;
			visu.stInteractiveError.xError := FALSE;
			uiState := 325;
		END_IF
		
		// Ignore
		IF visu.stInteractiveError.xBtnIgnore THEN
			visu.stInteractiveError.xBtnIgnore := FALSE;
			visu.stInteractiveError.xError := FALSE;
			uiState := visu.stInteractiveError.uiIgnoreState;
		END_IF
		
		// Abort
		IF visu.stInteractiveError.xBtnAbort THEN
			visu.stInteractiveError.xBtnAbort := FALSE;
			visu.stInteractiveError.xError := FALSE;
			uiState := visu.stInteractiveError.uiAbortState;
		END_IF
		
		// Reject order
		IF visu.stInteractiveError.xBtnRejectOrder THEN
			visu.stInteractiveError.xBtnRejectOrder := FALSE;
			visu.stInteractiveError.xError := FALSE;
			uiState := 480;
		END_IF		
		
	340:// Operation finished
		uiErrNo := stAppState.uiReturnCode;
		IF stAppState.xError THEN
			uiErrNo := 1;
		END_IF
		
		mesMES.OpEnd(udiONo := udiONo, uiOPos := uiOPos, uiCarrierId := uiCarrierId, uiErrNo := uiErrNo, pRcvHeader := ADR(stRcvHeader));
	
		uiState := 350;
		
	350:// Wait for MES request
		IF stRcvHeader.xDone THEN
			udiONo := strcvHeader.udiONo;
		    uiOPos := strcvHeader.uiOPos;
		    uiOpNo := strcvHeader.uiOpNo;
			uiState := 400;
		END_IF
		
	400:// Write RFID Data
		stRfidData.stMesData.udiONo := udiONo;
		stRfidData.stMesData.uiOPos := uiOPos;
		stRfidData.stMesData.uiOpNo := uiOpNo;
		stRfidData.stMesData.udiPNo := stRcvHeader.udiPNo;
		stRfidData.stMesData.uiResourceId := stRcvHeader.uiResourceId;
		stpStopper.WriteRfid(stRfidData);
		uiState := 410;
		
	410:// RFID write OK?
		IF stpStopper.xReady AND NOT stpStopper.dtmRfid.xTimeout THEN
			uiState := 375;
		ELSIF stpStopper.xReady THEN
			uiState := 500;
		END_IF
		
	480:// Send OPReset
		mesMES.OpReset(udiONo := udiONo, uiOPos := uiOPos, pRcvHeader := ADR(stRcvHeader));
		uiState := 481;
		
	481:// Wait for MES request
		IF stRcvHeader.xDone THEN
			uiState := 500;
		END_IF
		
	375:// Next operation for this resource?
		IF uiResourceId = stRcvHeader.uiResourceId THEN
			uiState := 110;
		ELSE
			uiState := 500;
		END_IF
		
	500:// Pass carrier
		IF NOT xSemaIn THEN
			xSemaOut := TRUE;
			stpStopper.Release();
			uiState := 505;
		END_IF
		
	505:// Wait for release
		IF stpStopper.xReady THEN
			uiState := 10;
		END_IF
	
END_CASE
END_METHOD

METHOD PRIVATE _DefaultMode : BOOL
VAR_INPUT
END_VAR
CASE uiState OF
	0:	// Idle
		convConveyor.Stop();
		IF xAuto THEN
			uiState := 1;
		END_IF
		
	1:	// Init
		convConveyor.RunToRight(FALSE);
		uiState := 2;
		
	
	2:	// Wait for RFID
		IF stpStopper.xReady AND stpStopper.xConnected THEN
			uiState := 10;
		END_IF
		
	10:	// Wait until carrier at stopper
		IF stpStopper.xCarrierAvailable AND NOT xCycleEnd THEN
			uiState := 15;
		END_IF
		
	15:	// Check if RFID tag recognized
		IF stpStopper.dtmRfid.stState.xTagPresent THEN
			uiState := 20;
		ELSE
			uiState := 500;
		END_IF
		
	20:	// Read RFID
		stpStopper.ReadRfid(ADR(stRfidData));
		uiState := 25;
		
	25:	// Wait until read finished
		IF stpStopper.xReady THEN
			uiState := 30;
		END_IF
		
	30:	// App. ready and active?
		IF stAppState.xReady AND stAppSettings.xActive THEN
			uiState := 50;
		ELSE
			uiState := 500;
		END_IF
		
	50:	// check carrier init condition
		IF stAppSettings.xCarrierInit THEN
			uiCondIn := 0;
			uiCondOut := astTransitionTable[0].uiCondOut;
			uiState := 55;
		ELSE
			// TODO: "dbAppPar".Init.iCntAct := 0; ???
			uiState := 60;
		END_IF
		
	55:	// check if Application is enabled in init step
		uiCarrierInitNum := uiCarrierInitNum + 1;
		IF uiCarrierInitNum >= stAppSettings.uiCarrierInitNum THEN
			uiCarrierInitNum := 0;
			stAppSettings.xCarrierInit := FALSE;
		END_IF	
	
		IF astTransitionTable[0].xAppEn THEN
			
			// Check if Application is active
			IF stAppSettings.xActive AND stAppState.xReady THEN
				uiActualTransitionRow := 0;
				uiState := 300;
			ELSE
				uiState := 490;
			END_IF
			
		ELSE
			
			SysMemSet(pDest := ADR(stRfidData.stMesData), udiValue := 0, udiCount := SIZEOF(stRfidData.stMesData));
			stRfidData.uiCode := astTransitionTable[0].uiCondOut;
			// TODO: "dbAppPar".Init.iCntAct := "dbAppPar".Init.iCntAct + 1;
			uiState := 400;
			
		END_IF
		
	60:	// Check if application is active
		IF stAppSettings.xActive THEN
			uiState := 65;
		ELSE
			uiState := 490;
		END_IF

	65:	// Check application start condition
        uiNextState := 490;
		
		// Search for a raw with the input condition
		uiCondIn := stRfidData.uiCode;
		uiCondOut := 0;
        FOR uiI := 1 TO 10 DO
            IF (uiCondIn = astTransitionTable[uiI].uiCondIn) AND (stRfidData.uiCode <> 0) THEN
				//Entry condition o.k.
                IF astTransitionTable[uiI].xAppEn THEN
                    // application for this condition activated
					uiActualTransitionRow := uiI;
					uiCondOut := astTransitionTable[uiI].uiCondOut;
                    uiNextState := 300;
                    EXIT;
                ELSE
                    // no application start, only write output code to RFID
                    stRfidData.uiCode := astTransitionTable[uiI].uiCondOut;
                    uiNextState := 400;
                    EXIT;
                END_IF
            END_IF
        END_FOR
		
        uiState := uiNextState;
		
	300:// Wait app. free
		IF stAppSettings.xActive AND stAppState.xReady THEN
			uiState := 305;
		END_IF
		
	305:// Send parameters to app
		stAppControl.uiOpNo := astTransitionTable[uiActualTransitionRow].uiPar1;
		SysMemCpy(pDest := ADR(stAppControl.auiPar), pSrc := ADR(astTransitionTable[uiActualTransitionRow].uiPar1), udiCount := 3 * SIZEOF(astTransitionTable[uiActualTransitionRow].uiPar1));
		uiState := 325;
		
	325:// Trigger App. start
		IF stAppSettings.xStopBelt THEN
			convConveyor.Stop();
		END_IF
		stAppControl.xStart := TRUE;
		uiState := 328;
		
	328:// Wait for App. started	
		IF NOT stAppState.xReady THEN
			stAppControl.xStart := FALSE;
			uiState := 330;
		END_IF
		
	330:// Wait for App. finished
		IF stAppState.xReady THEN
			convConveyor.RunToRight(FALSE);
			uiState := 335;
		END_IF
		
	335:// App. fininshed without error?
		IF stAppState.uiReturnCode = 0 THEN
			stRfidData.uiCode := astTransitionTable[uiActualTransitionRow].uiCondOut;
			uiState := 400;
		ELSE
			uiState := 336;
		END_IF
		
	336:// Interactive message
		Visu.stInteractiveError.xError := TRUE;
		Visu.stInteractiveError.sMessageID := UINT_TO_STRING(stAppState.uiReturnCode);
		visu.stInteractiveError.uiAbortState := 400;
		visu.stInteractiveError.uiIgnoreState := 400;
		
		// Retry
		IF visu.stInteractiveError.xBtnRepeat THEN
			visu.stInteractiveError.xBtnRepeat := FALSE;
			visu.stInteractiveError.xError := FALSE;
			uiState := 325;
		END_IF
		
		// Ignore
		IF visu.stInteractiveError.xBtnIgnore THEN
			visu.stInteractiveError.xBtnIgnore := FALSE;
			visu.stInteractiveError.xError := FALSE;
			uiState := visu.stInteractiveError.uiIgnoreState;
		END_IF
		
		// Abort
		IF visu.stInteractiveError.xBtnAbort THEN
			visu.stInteractiveError.xBtnAbort := FALSE;
			visu.stInteractiveError.xError := FALSE;
			uiState := visu.stInteractiveError.uiAbortState;
		END_IF		
		
	400:// Write RFID Data
		stpStopper.WriteRfid(stRfidData);
		uiState := 410;
		
	410:// Wait RFID write finished
		IF stpStopper.xReady THEN
			uiState := 500;
		END_IF
		
	490:// TODO
		// "dbVar".Hmi.StateCode[#iStNo].iOut := "dbVar".Hmi.StateCode[#iStNo].iIn; ???
		uiState := 500;	
		
	500:// Pass carrier
		IF NOT xSemaIn THEN
			xSemaOut := TRUE;
			stpStopper.Release();
			uiState := 505;
		END_IF
		
	505:// Wait for release
		IF stpStopper.xReady THEN
			uiState := 10;
		END_IF
	
END_CASE
END_METHOD

METHOD PRIVATE _ModuleCalls : BOOL
VAR_INPUT
END_VAR
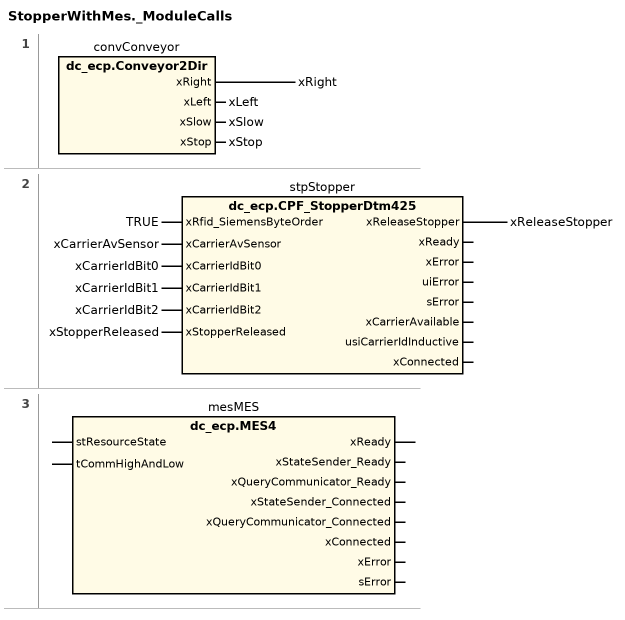
// NETWORK 1
convConveyor(xLeft => xLeft, xSlow => xSlow, xStop => xStop); // dc_ecp.Conveyor2Dir
xRight := convConveyor.xRight;

// NETWORK 2
stpStopper(
    xRfid_SiemensByteOrder := TRUE,
    xCarrierAvSensor := xCarrierAvSensor,
    xCarrierIdBit0 := xCarrierIdBit0,
    xCarrierIdBit1 := xCarrierIdBit1,
    xCarrierIdBit2 := xCarrierIdBit2,
    xStopperReleased := xStopperReleased); // dc_ecp.CPF_StopperDtm425
xReleaseStopper := stpStopper.xReleaseStopper;